      Contact( "CompALTA-MTA".FallaCompresor2 )
      wire#w4
      { S7_Templates := "SrcType := Int" } EQ_Contact(in1 := "DB-PrioridadesCmpAlta".Vcmp1, in2 := 2)
      wire#w5
      Contact( "DB-CompAltaDatos".Aut4 )
      Contact( "CompALTA-MTA".FallaCompresor4 )
      wire#w6
      { S7_Templates := "SrcType := Int" } EQ_Contact(in1 := "DB-PrioridadesCmpAlta".Vcmp4, in2 := 2)
   END_RUNG wire#w1
   RUNG wire#w4
      { S7_Templates := "SrcType := Int" } EQ_Contact(in1 := "DB-PrioridadesCmpAlta".Vcmp1, in2 := 1)
   END_RUNG wire#w5
   RUNG wire#w6
      { S7_Templates := "SrcType := Int" } EQ_Contact(in1 := "DB-PrioridadesCmpAlta".Vcmp4, in2 := 1)
   END_RUNG wire#w1
   RUNG wire#w5
      Contact( "DB-CompAltaDatos".Aut3 )
      Contact( "CompALTA-MTA".FallaCompresor3 )
      wire#w7
      { S7_Templates := "SrcType := Int" } EQ_Contact(in1 := "DB-PrioridadesCmpAlta".Vcmp3, in2 := 2)
   END_RUNG wire#w1
   RUNG wire#w7
      { S7_Templates := "SrcType := Int" } EQ_Contact(in1 := "DB-PrioridadesCmpAlta".Vcmp3, in2 := 1)
   END_RUNG wire#w1
   RUNG wire#w5
      Contact( "DB-CompAltaDatos".Aut2 )
      Contact( "CompALTA-MTA".FallaCompresor2 )
      wire#w8
      { S7_Templates := "SrcType := Int" } EQ_Contact(in1 := "DB-PrioridadesCmpAlta".Vcmp2, in2 := 2)
   END_RUNG wire#w1
   RUNG wire#w8
      { S7_Templates := "SrcType := Int" } EQ_Contact(in1 := "DB-PrioridadesCmpAlta".Vcmp2, in2 := 1)
   END_RUNG wire#w1
   RUNG wire#w3
      Contact( "DB-CompAltaDatos".Aut2 )
      Contact( "CompALTA-MTA".FallaCompresor2 )
      wire#w9
      { S7_Templates := "SrcType := Int" } EQ_Contact(in1 := "DB-PrioridadesCmpAlta".Vcmp2, in2 := 2)
      wire#w10
      Contact( "DB-CompAltaDatos".Aut4 )
      Contact( "CompALTA-MTA".FallaCompresor4 )
      wire#w11
      { S7_Templates := "SrcType := Int" } EQ_Contact(in1 := "DB-PrioridadesCmpAlta".Vcmp4, in2 := 2)
   END_RUNG wire#w1
   RUNG wire#w9
      { S7_Templates := "SrcType := Int" } EQ_Contact(in1 := "DB-PrioridadesCmpAlta".Vcmp2, in2 := 1)
   END_RUNG wire#w10
   RUNG wire#w11
      { S7_Templates := "SrcType := Int" } EQ_Contact(in1 := "DB-PrioridadesCmpAlta".Vcmp4, in2 := 1)
   END_RUNG wire#w1
   RUNG wire#w10
      Contact( "DB-CompAltaDatos".Aut3 )
      Contact( "CompALTA-MTA".FallaCompresor3 )
      wire#w12
      { S7_Templates := "SrcType := Int" } EQ_Contact(in1 := "DB-PrioridadesCmpAlta".Vcmp3, in2 := 2)
   END_RUNG wire#w1
   RUNG wire#w12
      { S7_Templates := "SrcType := Int" } EQ_Contact(in1 := "DB-PrioridadesCmpAlta".Vcmp3, in2 := 1)
   END_RUNG wire#w1
   RUNG wire#w3
      Contact( "DB-CompAltaDatos".Aut3 )
      Contact( "CompALTA-MTA".FallaCompresor3 )
      wire#w13
      { S7_Templates := "SrcType := Int" } EQ_Contact(in1 := "DB-PrioridadesCmpAlta".Vcmp3, in2 := 2)
      wire#w14
      Contact( "DB-CompAltaDatos".Aut4 )
      Contact( "CompALTA-MTA".FallaCompresor4 )
      wire#w15
      { S7_Templates := "SrcType := Int" } EQ_Contact(in1 := "DB-PrioridadesCmpAlta".Vcmp4, in2 := 2)
   END_RUNG wire#w1
   RUNG wire#w13
      { S7_Templates := "SrcType := Int" } EQ_Contact(in1 := "DB-PrioridadesCmpAlta".Vcmp3, in2 := 1)
   END_RUNG wire#w14
   RUNG wire#w15
      { S7_Templates := "SrcType := Int" } EQ_Contact(in1 := "DB-PrioridadesCmpAlta".Vcmp4, in2 := 1)
   END_RUNG wire#w1
   RUNG wire#powerrail
      { S7_Templates := "SrcType := Int" } EQ_Contact(in1 := "DB-PrioridadesCmpAlta".Vcmp5, in2 := 4)
      wire#w16
      Contact( "DB-CompAltaDatos".Aut1 )
      Contact( "CompALTA-MTA".FallaCompresor1 )
      wire#w17
      { S7_Templates := "SrcType := Int" } EQ_Contact(in1 := "DB-PrioridadesCmpAlta".Vcmp1, in2 := 3)
      wire#w18
      Contact( "DB-CompAltaDatos".Aut4 )
      Contact( "CompALTA-MTA".FallaCompresor4 )
      wire#w19
      { S7_Templates := "SrcType := Int" } EQ_Contact(in1 := "DB-PrioridadesCmpAlta".Vcmp4, in2 := 3)
      wire#w20
      Contact( "DB-CompAltaDatos".Aut2 )
      Contact( "CompALTA-MTA".FallaCompresor2 )
      wire#w21
      { S7_Templates := "SrcType := Int" } EQ_Contact(in1 := "DB-PrioridadesCmpAlta".Vcmp2, in2 := 3)
   END_RUNG wire#w1
   RUNG wire#w17
      { S7_Templates := "SrcType := Int" } EQ_Contact(in1 := "DB-PrioridadesCmpAlta".Vcmp1, in2 := 2)
   END_RUNG wire#w18
   RUNG wire#w17
      { S7_Templates := "SrcType := Int" } EQ_Contact(in1 := "DB-PrioridadesCmpAlta".Vcmp1, in2 := 1)
   END_RUNG wire#w18
   RUNG wire#w19
      { S7_Templates := "SrcType := Int" } EQ_Contact(in1 := "DB-PrioridadesCmpAlta".Vcmp4, in2 := 2)
   END_RUNG wire#w20
   RUNG wire#w19
      { S7_Templates := "SrcType := Int" } EQ_Contact(in1 := "DB-PrioridadesCmpAlta".Vcmp4, in2 := 1)
   END_RUNG wire#w20
   RUNG wire#w21
      { S7_Templates := "SrcType := Int" } EQ_Contact(in1 := "DB-PrioridadesCmpAlta".Vcmp2, in2 := 2)
   END_RUNG wire#w1
   RUNG wire#w21
      { S7_Templates := "SrcType := Int" } EQ_Contact(in1 := "DB-PrioridadesCmpAlta".Vcmp2, in2 := 1)
   END_RUNG wire#w1
   RUNG wire#w20
      Contact( "DB-CompAltaDatos".Aut4 )
      Contact( "CompALTA-MTA".FallaCompresor4 )
      wire#w22
      { S7_Templates := "SrcType := Int" } EQ_Contact(in1 := "DB-PrioridadesCmpAlta".Vcmp4, in2 := 3)
   END_RUNG wire#w1
   RUNG wire#w22
      { S7_Templates := "SrcType := Int" } EQ_Contact(in1 := "DB-PrioridadesCmpAlta".Vcmp4, in2 := 2)
   END_RUNG wire#w1
   RUNG wire#w22
      { S7_Templates := "SrcType := Int" } EQ_Contact(in1 := "DB-PrioridadesCmpAlta".Vcmp4, in2 := 1)
   END_RUNG wire#w1
   RUNG wire#w18
      Contact( "DB-CompAltaDatos".Aut3 )
      Contact( "CompALTA-MTA".FallaCompresor3 )
      wire#w23
      { S7_Templates := "SrcType := Int" } EQ_Contact(in1 := "DB-PrioridadesCmpAlta".Vcmp3, in2 := 3)
      wire#w24
      Contact( "DB-CompAltaDatos".Aut2 )
      Contact( "CompALTA-MTA".FallaCompresor2 )
      wire#w25
      { S7_Templates := "SrcType := Int" } EQ_Contact(in1 := "DB-PrioridadesCmpAlta".Vcmp2, in2 := 3)
   END_RUNG wire#w1
   RUNG wire#w23
      { S7_Templates := "SrcType := Int" } EQ_Contact(in1 := "DB-PrioridadesCmpAlta".Vcmp3, in2 := 2)
   END_RUNG wire#w24
   RUNG wire#w23
      { S7_Templates := "SrcType := Int" } EQ_Contact(in1 := "DB-PrioridadesCmpAlta".Vcmp3, in2 := 1)
   END_RUNG wire#w24
   RUNG wire#w25
      { S7_Templates := "SrcType := Int" } EQ_Contact(in1 := "DB-PrioridadesCmpAlta".Vcmp2, in2 := 2)
   END_RUNG wire#w1
   RUNG wire#w25
      { S7_Templates := "SrcType := Int" } EQ_Contact(in1 := "DB-PrioridadesCmpAlta".Vcmp2, in2 := 1)
   END_RUNG wire#w1
   RUNG wire#w16
      Contact( "DB-CompAltaDatos".Aut2 )
      Contact( "CompALTA-MTA".FallaCompresor2 )
      wire#w26
      { S7_Templates := "SrcType := Int" } EQ_Contact(in1 := "DB-PrioridadesCmpAlta".Vcmp2, in2 := 3)
      wire#w27
      Contact( "DB-CompAltaDatos".Aut4 )
      Contact( "CompALTA-MTA".FallaCompresor4 )
      wire#w28
      { S7_Templates := "SrcType := Int" } EQ_Contact(in1 := "DB-PrioridadesCmpAlta".Vcmp4, in2 := 3)
      wire#w29
      Contact( "DB-CompAltaDatos".Aut3 )
      Contact( "CompALTA-MTA".FallaCompresor3 )
      wire#w30
      { S7_Templates := "SrcType := Int" } EQ_Contact(in1 := "DB-PrioridadesCmpAlta".Vcmp3, in2 := 3)
   END_RUNG wire#w1
   RUNG wire#w26
      { S7_Templates := "SrcType := Int" } EQ_Contact(in1 := "DB-PrioridadesCmpAlta".Vcmp2, in2 := 2)
   END_RUNG wire#w27
   RUNG wire#w26
      { S7_Templates := "SrcType := Int" } EQ_Contact(in1 := "DB-PrioridadesCmpAlta".Vcmp2, in2 := 1)
   END_RUNG wire#w27
   RUNG wire#w28
      { S7_Templates := "SrcType := Int" } EQ_Contact(in1 := "DB-PrioridadesCmpAlta".Vcmp4, in2 := 2)
   END_RUNG wire#w29
   RUNG wire#w28
      { S7_Templates := "SrcType := Int" } EQ_Contact(in1 := "DB-PrioridadesCmpAlta".Vcmp4, in2 := 1)
   END_RUNG wire#w29
   RUNG wire#w30
      { S7_Templates := "SrcType := Int" } EQ_Contact(in1 := "DB-PrioridadesCmpAlta".Vcmp3, in2 := 2)
   END_RUNG wire#w1
   RUNG wire#w30
      { S7_Templates := "SrcType := Int" } EQ_Contact(in1 := "DB-PrioridadesCmpAlta".Vcmp3, in2 := 1)
   END_RUNG wire#w1
   RUNG wire#powerrail
      { S7_Templates := "SrcType := Int" } EQ_Contact(in1 := "DB-PrioridadesCmpAlta".Vcmp5, in2 := 5)
      Contact( "DB-CompAltaDatos".Aut1 )
      Contact( "CompALTA-MTA".FallaCompresor1 )
      Contact( "DB-CompAltaDatos".Aut2 )
      Contact( "CompALTA-MTA".FallaCompresor2 )
      Contact( "DB-CompAltaDatos".Aut3 )
      Contact( "CompALTA-MTA".FallaCompresor3 )
      Contact( "DB-CompAltaDatos".Aut4 )
      Contact( "CompALTA-MTA".FallaCompresor4 )
   END_RUNG wire#w1
   // the same network as SCL:
   IF (("DB-PrioridadesCmpAlta".Vcmp5 = 1) OR (("DB-PrioridadesCmpAlta".Vcmp5 = 2) AND (("DB-CompAltaDatos".Aut1 AND "CompALTA-MTA".FallaCompresor1 AND ("DB-PrioridadesCmpAlta".Vcmp1 = 1)) OR ("DB-CompAltaDatos".Aut2 AND "CompALTA-MTA".FallaCompresor2 AND ("DB-PrioridadesCmpAlta".Vcmp2 = 1)) OR ("DB-CompAltaDatos".Aut3 AND "CompALTA-MTA".FallaCompresor3 AND ("DB-PrioridadesCmpAlta".Vcmp3 = 1)) OR ("DB-CompAltaDatos".Aut4 AND "CompALTA-MTA".FallaCompresor4 AND ("DB-PrioridadesCmpAlta".Vcmp4 = 1)))) OR (("DB-PrioridadesCmpAlta".Vcmp5 = 3) AND (("DB-CompAltaDatos".Aut2 AND "CompALTA-MTA".FallaCompresor2 AND (("DB-PrioridadesCmpAlta".Vcmp1 = 2) OR ("DB-PrioridadesCmpAlta".Vcmp1 = 1)) AND (("DB-CompAltaDatos".Aut4 AND "CompALTA-MTA".FallaCompresor4 AND (("DB-PrioridadesCmpAlta".Vcmp4 = 2) OR ("DB-PrioridadesCmpAlta".Vcmp4 = 1))) OR ("DB-CompAltaDatos".Aut3 AND "CompALTA-MTA".FallaCompresor3 AND (("DB-PrioridadesCmpAlta".Vcmp3 = 2) OR ("DB-PrioridadesCmpAlta".Vcmp3 = 1))) OR ("DB-CompAltaDatos".Aut2 AND "CompALTA-MTA".FallaCompresor2 AND (("DB-PrioridadesCmpAlta".Vcmp2 = 2) OR ("DB-PrioridadesCmpAlta".Vcmp2 = 1))))) OR ("DB-CompAltaDatos".Aut2 AND "CompALTA-MTA".FallaCompresor2 AND (("DB-PrioridadesCmpAlta".Vcmp2 = 2) OR ("DB-PrioridadesCmpAlta".Vcmp2 = 1)) AND (("DB-CompAltaDatos".Aut4 AND "CompALTA-MTA".FallaCompresor4 AND (("DB-PrioridadesCmpAlta".Vcmp4 = 2) OR ("DB-PrioridadesCmpAlta".Vcmp4 = 1))) OR ("DB-CompAltaDatos".Aut3 AND "CompALTA-MTA".FallaCompresor3 AND (("DB-PrioridadesCmpAlta".Vcmp3 = 2) OR ("DB-PrioridadesCmpAlta".Vcmp3 = 1))))) OR ("DB-CompAltaDatos".Aut3 AND "CompALTA-MTA".FallaCompresor3 AND (("DB-PrioridadesCmpAlta".Vcmp3 = 2) OR ("DB-PrioridadesCmpAlta".Vcmp3 = 1)) AND "DB-CompAltaDatos".Aut4 AND "CompALTA-MTA".FallaCompresor4 AND (("DB-PrioridadesCmpAlta".Vcmp4 = 2) OR ("DB-PrioridadesCmpAlta".Vcmp4 = 1))))) OR (("DB-PrioridadesCmpAlta".Vcmp5 = 4) AND (("DB-CompAltaDatos".Aut1 AND "CompALTA-MTA".FallaCompresor1 AND (("DB-PrioridadesCmpAlta".Vcmp1 = 3) OR ("DB-PrioridadesCmpAlta".Vcmp1 = 2) OR ("DB-PrioridadesCmpAlta".Vcmp1 = 1)) AND (("DB-CompAltaDatos".Aut4 AND "CompALTA-MTA".FallaCompresor4 AND (("DB-PrioridadesCmpAlta".Vcmp4 = 3) OR ("DB-PrioridadesCmpAlta".Vcmp4 = 2) OR ("DB-PrioridadesCmpAlta".Vcmp4 = 1)) AND (("DB-CompAltaDatos".Aut2 AND "CompALTA-MTA".FallaCompresor2 AND (("DB-PrioridadesCmpAlta".Vcmp2 = 3) OR ("DB-PrioridadesCmpAlta".Vcmp2 = 2) OR ("DB-PrioridadesCmpAlta".Vcmp2 = 1))) OR ("DB-CompAltaDatos".Aut4 AND "CompALTA-MTA".FallaCompresor4 AND (("DB-PrioridadesCmpAlta".Vcmp4 = 3) OR ("DB-PrioridadesCmpAlta".Vcmp4 = 2) OR ("DB-PrioridadesCmpAlta".Vcmp4 = 1))))) OR ("DB-CompAltaDatos".Aut3 AND "CompALTA-MTA".FallaCompresor3 AND (("DB-PrioridadesCmpAlta".Vcmp3 = 3) OR ("DB-PrioridadesCmpAlta".Vcmp3 = 2) OR ("DB-PrioridadesCmpAlta".Vcmp3 = 1)) AND "DB-CompAltaDatos".Aut2 AND "CompALTA-MTA".FallaCompresor2 AND (("DB-PrioridadesCmpAlta".Vcmp2 = 3) OR ("DB-PrioridadesCmpAlta".Vcmp2 = 2) OR ("DB-PrioridadesCmpAlta".Vcmp2 = 1))))) OR ("DB-CompAltaDatos".Aut2 AND "CompALTA-MTA".FallaCompresor2 AND (("DB-PrioridadesCmpAlta".Vcmp2 = 3) OR ("DB-PrioridadesCmpAlta".Vcmp2 = 2) OR ("DB-PrioridadesCmpAlta".Vcmp2 = 1)) AND "DB-CompAltaDatos".Aut4 AND "CompALTA-MTA".FallaCompresor4 AND (("DB-PrioridadesCmpAlta".Vcmp4 = 3) OR ("DB-PrioridadesCmpAlta".Vcmp4 = 2) OR ("DB-PrioridadesCmpAlta".Vcmp4 = 1)) AND "DB-CompAltaDatos".Aut3 AND "CompALTA-MTA".FallaCompresor3 AND (("DB-PrioridadesCmpAlta".Vcmp3 = 3) OR ("DB-PrioridadesCmpAlta".Vcmp3 = 2) OR ("DB-PrioridadesCmpAlta".Vcmp3 = 1))))) OR (("DB-PrioridadesCmpAlta".Vcmp5 = 5) AND "DB-CompAltaDatos".Aut1 AND "CompALTA-MTA".FallaCompresor1 AND "DB-CompAltaDatos".Aut2 AND "CompALTA-MTA".FallaCompresor2 AND "DB-CompAltaDatos".Aut3 AND "CompALTA-MTA".FallaCompresor3 AND "DB-CompAltaDatos".Aut4 AND "CompALTA-MTA".FallaCompresor4)) AND "DB-CompAltaDatos".Aut5 AND NOT "CompALTA-MTA".FallaCompresor5 THEN
       "CompALTA-MTA".VRealCmp5 := 1;
   END_IF;
END_REGION
END_FUNCTION

FUNCTION "FlancosCmpAlta" : Void   // FC45, LAD
{ S7_Optimized_Access := 'FALSE' }
VERSION : 0.1
   VAR_TEMP   // added for the SCL form of the ladder/FBD networks
      _w1 : Bool;
      _w2 : Bool;
      _w3 : Bool;
      _w4 : Bool;
      _w5 : Bool;
      _w6 : Bool;
      _w7 : Bool;
      _s5time1 : S5Time;
   END_VAR
BEGIN

REGION Network 1
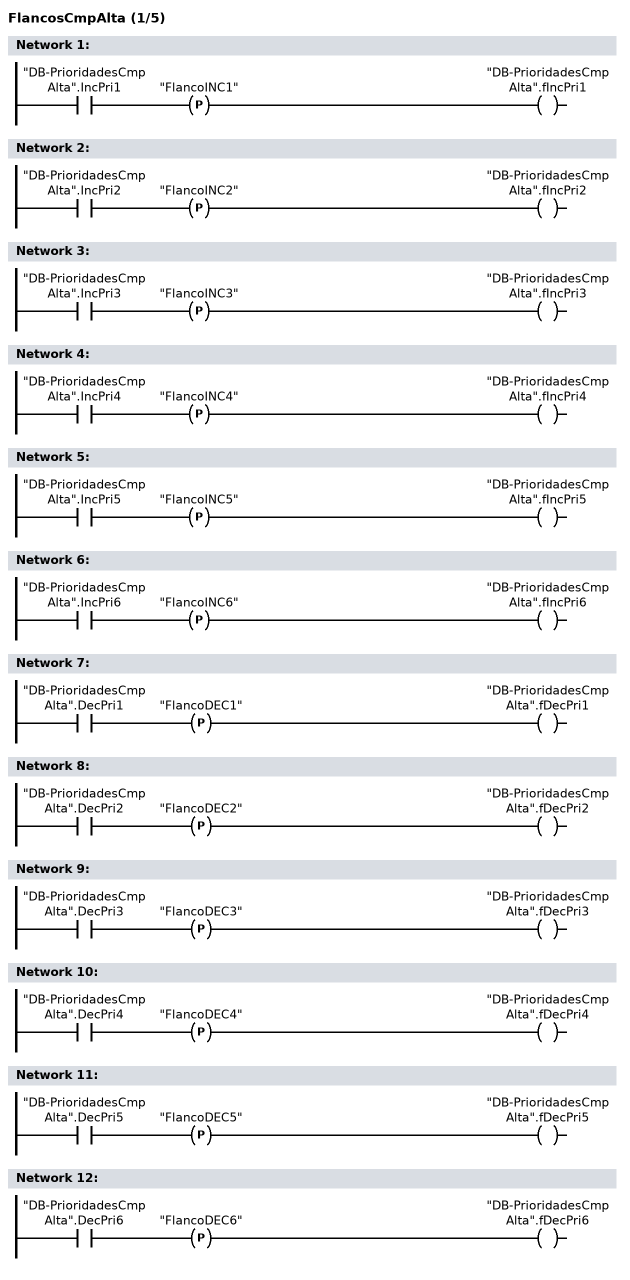
   RUNG wire#powerrail
      Contact( "DB-PrioridadesCmpAlta".IncPri1 )
      P_Trig( "FlancoINC1" )
      Coil( "DB-PrioridadesCmpAlta".fIncPri1 )
   END_RUNG
   // the same network as SCL:
   #_w1 := "DB-PrioridadesCmpAlta".IncPri1 AND NOT "FlancoINC1";   // rising edge
   "FlancoINC1" := "DB-PrioridadesCmpAlta".IncPri1;
   "DB-PrioridadesCmpAlta".fIncPri1 := #_w1;
END_REGION

REGION Network 2
   RUNG wire#powerrail
      Contact( "DB-PrioridadesCmpAlta".IncPri2 )
      P_Trig( "FlancoINC2" )
      Coil( "DB-PrioridadesCmpAlta".fIncPri2 )
   END_RUNG
   // the same network as SCL:
   #_w1 := "DB-PrioridadesCmpAlta".IncPri2 AND NOT "FlancoINC2";   // rising edge
   "FlancoINC2" := "DB-PrioridadesCmpAlta".IncPri2;
   "DB-PrioridadesCmpAlta".fIncPri2 := #_w1;
END_REGION

REGION Network 3
   RUNG wire#powerrail
      Contact( "DB-PrioridadesCmpAlta".IncPri3 )
      P_Trig( "FlancoINC3" )
      Coil( "DB-PrioridadesCmpAlta".fIncPri3 )
   END_RUNG
   // the same network as SCL:
   #_w1 := "DB-PrioridadesCmpAlta".IncPri3 AND NOT "FlancoINC3";   // rising edge
   "FlancoINC3" := "DB-PrioridadesCmpAlta".IncPri3;
   "DB-PrioridadesCmpAlta".fIncPri3 := #_w1;
END_REGION

REGION Network 4
   RUNG wire#powerrail
      Contact( "DB-PrioridadesCmpAlta".IncPri4 )
      P_Trig( "FlancoINC4" )
      Coil( "DB-PrioridadesCmpAlta".fIncPri4 )
   END_RUNG
   // the same network as SCL:
   #_w1 := "DB-PrioridadesCmpAlta".IncPri4 AND NOT "FlancoINC4";   // rising edge
   "FlancoINC4" := "DB-PrioridadesCmpAlta".IncPri4;
   "DB-PrioridadesCmpAlta".fIncPri4 := #_w1;
END_REGION

REGION Network 5
   RUNG wire#powerrail
      Contact( "DB-PrioridadesCmpAlta".IncPri5 )
      P_Trig( "FlancoINC5" )
      Coil( "DB-PrioridadesCmpAlta".fIncPri5 )
   END_RUNG
   // the same network as SCL:
   #_w1 := "DB-PrioridadesCmpAlta".IncPri5 AND NOT "FlancoINC5";   // rising edge
   "FlancoINC5" := "DB-PrioridadesCmpAlta".IncPri5;
   "DB-PrioridadesCmpAlta".fIncPri5 := #_w1;
END_REGION

REGION Network 6
   RUNG wire#powerrail
      Contact( "DB-PrioridadesCmpAlta".IncPri6 )
      P_Trig( "FlancoINC6" )
      Coil( "DB-PrioridadesCmpAlta".fIncPri6 )
   END_RUNG
   // the same network as SCL:
   #_w1 := "DB-PrioridadesCmpAlta".IncPri6 AND NOT "FlancoINC6";   // rising edge
   "FlancoINC6" := "DB-PrioridadesCmpAlta".IncPri6;
   "DB-PrioridadesCmpAlta".fIncPri6 := #_w1;
END_REGION

REGION Network 7
   RUNG wire#powerrail
      Contact( "DB-PrioridadesCmpAlta".DecPri1 )
      P_Trig( "FlancoDEC1" )
      Coil( "DB-PrioridadesCmpAlta".fDecPri1 )
   END_RUNG
   // the same network as SCL:
   #_w1 := "DB-PrioridadesCmpAlta".DecPri1 AND NOT "FlancoDEC1";   // rising edge
   "FlancoDEC1" := "DB-PrioridadesCmpAlta".DecPri1;
   "DB-PrioridadesCmpAlta".fDecPri1 := #_w1;
END_REGION

REGION Network 8
   RUNG wire#powerrail
      Contact( "DB-PrioridadesCmpAlta".DecPri2 )
      P_Trig( "FlancoDEC2" )
      Coil( "DB-PrioridadesCmpAlta".fDecPri2 )
   END_RUNG
   // the same network as SCL:
   #_w1 := "DB-PrioridadesCmpAlta".DecPri2 AND NOT "FlancoDEC2";   // rising edge
   "FlancoDEC2" := "DB-PrioridadesCmpAlta".DecPri2;
   "DB-PrioridadesCmpAlta".fDecPri2 := #_w1;
END_REGION

REGION Network 9
   RUNG wire#powerrail
      Contact( "DB-PrioridadesCmpAlta".DecPri3 )
      P_Trig( "FlancoDEC3" )
      Coil( "DB-PrioridadesCmpAlta".fDecPri3 )
   END_RUNG
   // the same network as SCL:
   #_w1 := "DB-PrioridadesCmpAlta".DecPri3 AND NOT "FlancoDEC3";   // rising edge
   "FlancoDEC3" := "DB-PrioridadesCmpAlta".DecPri3;
   "DB-PrioridadesCmpAlta".fDecPri3 := #_w1;
END_REGION

REGION Network 10
   RUNG wire#powerrail
      Contact( "DB-PrioridadesCmpAlta".DecPri4 )
      P_Trig( "FlancoDEC4" )
      Coil( "DB-PrioridadesCmpAlta".fDecPri4 )
   END_RUNG
   // the same network as SCL:
   #_w1 := "DB-PrioridadesCmpAlta".DecPri4 AND NOT "FlancoDEC4";   // rising edge
   "FlancoDEC4" := "DB-PrioridadesCmpAlta".DecPri4;
   "DB-PrioridadesCmpAlta".fDecPri4 := #_w1;
END_REGION

REGION Network 11
   RUNG wire#powerrail
      Contact( "DB-PrioridadesCmpAlta".DecPri5 )
      P_Trig( "FlancoDEC5" )
      Coil( "DB-PrioridadesCmpAlta".fDecPri5 )
   END_RUNG
   // the same network as SCL:
   #_w1 := "DB-PrioridadesCmpAlta".DecPri5 AND NOT "FlancoDEC5";   // rising edge
   "FlancoDEC5" := "DB-PrioridadesCmpAlta".DecPri5;
   "DB-PrioridadesCmpAlta".fDecPri5 := #_w1;
END_REGION

REGION Network 12
   RUNG wire#powerrail
      Contact( "DB-PrioridadesCmpAlta".DecPri6 )
      P_Trig( "FlancoDEC6" )
      Coil( "DB-PrioridadesCmpAlta".fDecPri6 )
   END_RUNG
   // the same network as SCL:
   #_w1 := "DB-PrioridadesCmpAlta".DecPri6 AND NOT "FlancoDEC6";   // rising edge
   "FlancoDEC6" := "DB-PrioridadesCmpAlta".DecPri6;
   "DB-PrioridadesCmpAlta".fDecPri6 := #_w1;
END_REGION

REGION Network 13
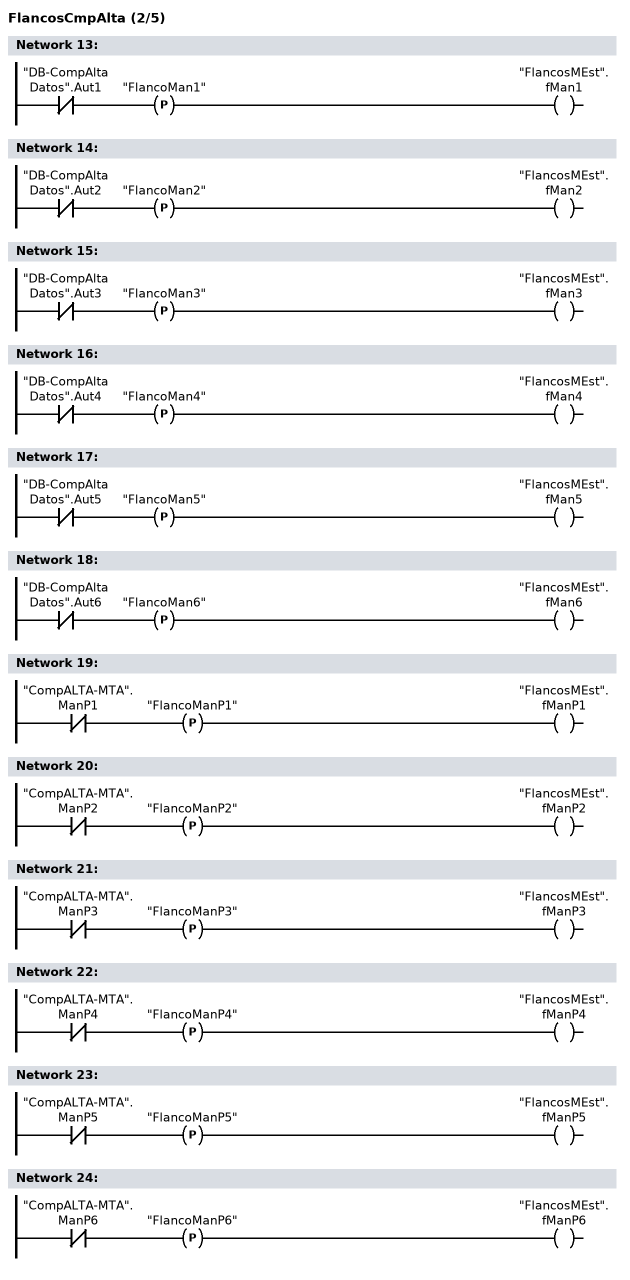
   RUNG wire#powerrail
      I_Contact( "DB-CompAltaDatos".Aut1 )
      P_Trig( "FlancoMan1" )
      Coil( "FlancosMEst".fMan1 )
   END_RUNG
   // the same network as SCL:
   #_w1 := NOT "DB-CompAltaDatos".Aut1 AND NOT "FlancoMan1";   // rising edge
   "FlancoMan1" := NOT "DB-CompAltaDatos".Aut1;
   "FlancosMEst".fMan1 := #_w1;
END_REGION

REGION Network 14
   RUNG wire#powerrail
      I_Contact( "DB-CompAltaDatos".Aut2 )
      P_Trig( "FlancoMan2" )
      Coil( "FlancosMEst".fMan2 )
   END_RUNG
   // the same network as SCL:
   #_w1 := NOT "DB-CompAltaDatos".Aut2 AND NOT "FlancoMan2";   // rising edge
   "FlancoMan2" := NOT "DB-CompAltaDatos".Aut2;
   "FlancosMEst".fMan2 := #_w1;
END_REGION

REGION Network 15
   RUNG wire#powerrail
      I_Contact( "DB-CompAltaDatos".Aut3 )
      P_Trig( "FlancoMan3" )
      Coil( "FlancosMEst".fMan3 )
   END_RUNG
   // the same network as SCL:
   #_w1 := NOT "DB-CompAltaDatos".Aut3 AND NOT "FlancoMan3";   // rising edge
   "FlancoMan3" := NOT "DB-CompAltaDatos".Aut3;
   "FlancosMEst".fMan3 := #_w1;
END_REGION

REGION Network 16
   RUNG wire#powerrail
      I_Contact( "DB-CompAltaDatos".Aut4 )
      P_Trig( "FlancoMan4" )
      Coil( "FlancosMEst".fMan4 )
   END_RUNG
   // the same network as SCL:
   #_w1 := NOT "DB-CompAltaDatos".Aut4 AND NOT "FlancoMan4";   // rising edge
   "FlancoMan4" := NOT "DB-CompAltaDatos".Aut4;
   "FlancosMEst".fMan4 := #_w1;
END_REGION

REGION Network 17
   RUNG wire#powerrail
      I_Contact( "DB-CompAltaDatos".Aut5 )
      P_Trig( "FlancoMan5" )
      Coil( "FlancosMEst".fMan5 )
   END_RUNG
   // the same network as SCL:
   #_w1 := NOT "DB-CompAltaDatos".Aut5 AND NOT "FlancoMan5";   // rising edge
   "FlancoMan5" := NOT "DB-CompAltaDatos".Aut5;
   "FlancosMEst".fMan5 := #_w1;
END_REGION

REGION Network 18
   RUNG wire#powerrail
      I_Contact( "DB-CompAltaDatos".Aut6 )
      P_Trig( "FlancoMan6" )
      Coil( "FlancosMEst".fMan6 )
   END_RUNG
   // the same network as SCL:
   #_w1 := NOT "DB-CompAltaDatos".Aut6 AND NOT "FlancoMan6";   // rising edge
   "FlancoMan6" := NOT "DB-CompAltaDatos".Aut6;
   "FlancosMEst".fMan6 := #_w1;
END_REGION

REGION Network 19
   RUNG wire#powerrail
      I_Contact( "CompALTA-MTA".ManP1 )
      P_Trig( "FlancoManP1" )
      Coil( "FlancosMEst".fManP1 )
   END_RUNG
   // the same network as SCL:
   #_w1 := NOT "CompALTA-MTA".ManP1 AND NOT "FlancoManP1";   // rising edge
   "FlancoManP1" := NOT "CompALTA-MTA".ManP1;
   "FlancosMEst".fManP1 := #_w1;
END_REGION

REGION Network 20
   RUNG wire#powerrail
      I_Contact( "CompALTA-MTA".ManP2 )
      P_Trig( "FlancoManP2" )
      Coil( "FlancosMEst".fManP2 )
   END_RUNG
   // the same network as SCL:
   #_w1 := NOT "CompALTA-MTA".ManP2 AND NOT "FlancoManP2";   // rising edge
   "FlancoManP2" := NOT "CompALTA-MTA".ManP2;
   "FlancosMEst".fManP2 := #_w1;
END_REGION

REGION Network 21
   RUNG wire#powerrail
      I_Contact( "CompALTA-MTA".ManP3 )
      P_Trig( "FlancoManP3" )
      Coil( "FlancosMEst".fManP3 )
   END_RUNG
   // the same network as SCL:
   #_w1 := NOT "CompALTA-MTA".ManP3 AND NOT "FlancoManP3";   // rising edge
   "FlancoManP3" := NOT "CompALTA-MTA".ManP3;
   "FlancosMEst".fManP3 := #_w1;
END_REGION

REGION Network 22
   RUNG wire#powerrail
      I_Contact( "CompALTA-MTA".ManP4 )
      P_Trig( "FlancoManP4" )
      Coil( "FlancosMEst".fManP4 )
   END_RUNG
   // the same network as SCL:
   #_w1 := NOT "CompALTA-MTA".ManP4 AND NOT "FlancoManP4";   // rising edge
   "FlancoManP4" := NOT "CompALTA-MTA".ManP4;
   "FlancosMEst".fManP4 := #_w1;
END_REGION

REGION Network 23
   RUNG wire#powerrail
      I_Contact( "CompALTA-MTA".ManP5 )
      P_Trig( "FlancoManP5" )
      Coil( "FlancosMEst".fManP5 )
   END_RUNG
   // the same network as SCL:
   #_w1 := NOT "CompALTA-MTA".ManP5 AND NOT "FlancoManP5";   // rising edge
   "FlancoManP5" := NOT "CompALTA-MTA".ManP5;
   "FlancosMEst".fManP5 := #_w1;
END_REGION

REGION Network 24
   RUNG wire#powerrail
      I_Contact( "CompALTA-MTA".ManP6 )
      P_Trig( "FlancoManP6" )
      Coil( "FlancosMEst".fManP6 )
   END_RUNG
   // the same network as SCL:
   #_w1 := NOT "CompALTA-MTA".ManP6 AND NOT "FlancoManP6";   // rising edge
   "FlancoManP6" := NOT "CompALTA-MTA".ManP6;
   "FlancosMEst".fManP6 := #_w1;
END_REGION

REGION Network 25
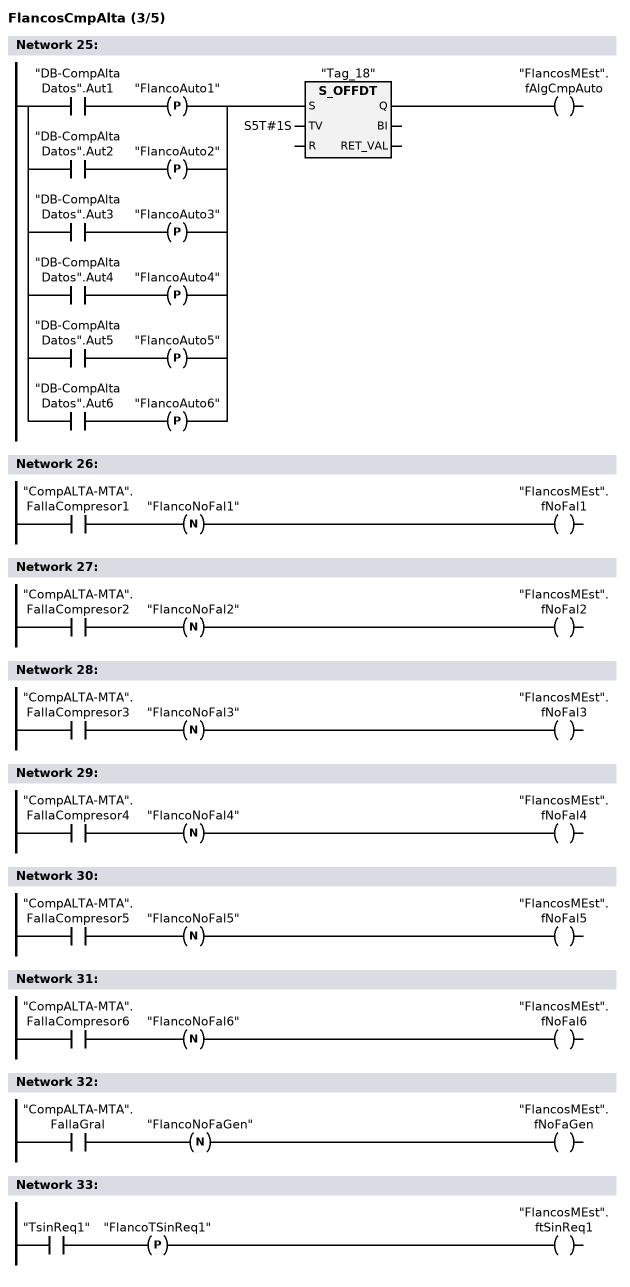
   RUNG wire#powerrail
      Contact( "DB-CompAltaDatos".Aut1 )
      P_Trig( "FlancoAuto1" )
      wire#w1
      S_OFFDT(T_NO := "Tag_18", TV := S5T#1S, R :=, BI =>, RET_VAL =>)
      Coil( "FlancosMEst".fAlgCmpAuto )
   END_RUNG
   RUNG wire#powerrail
      Contact( "DB-CompAltaDatos".Aut2 )
      P_Trig( "FlancoAuto2" )
   END_RUNG wire#w1
   RUNG wire#powerrail
      Contact( "DB-CompAltaDatos".Aut3 )
      P_Trig( "FlancoAuto3" )
   END_RUNG wire#w1
   RUNG wire#powerrail
      Contact( "DB-CompAltaDatos".Aut4 )
      P_Trig( "FlancoAuto4" )
   END_RUNG wire#w1
   RUNG wire#powerrail
      Contact( "DB-CompAltaDatos".Aut5 )
      P_Trig( "FlancoAuto5" )
   END_RUNG wire#w1
   RUNG wire#powerrail
      Contact( "DB-CompAltaDatos".Aut6 )
      P_Trig( "FlancoAuto6" )
   END_RUNG wire#w1
   // the same network as SCL:
   #_w1 := "DB-CompAltaDatos".Aut1 AND NOT "FlancoAuto1";   // rising edge
   "FlancoAuto1" := "DB-CompAltaDatos".Aut1;
   #_w2 := "DB-CompAltaDatos".Aut2 AND NOT "FlancoAuto2";   // rising edge
   "FlancoAuto2" := "DB-CompAltaDatos".Aut2;
   #_w3 := "DB-CompAltaDatos".Aut3 AND NOT "FlancoAuto3";   // rising edge
   "FlancoAuto3" := "DB-CompAltaDatos".Aut3;
   #_w4 := "DB-CompAltaDatos".Aut4 AND NOT "FlancoAuto4";   // rising edge
   "FlancoAuto4" := "DB-CompAltaDatos".Aut4;
   #_w5 := "DB-CompAltaDatos".Aut5 AND NOT "FlancoAuto5";   // rising edge
   "FlancoAuto5" := "DB-CompAltaDatos".Aut5;
   #_w6 := "DB-CompAltaDatos".Aut6 AND NOT "FlancoAuto6";   // rising edge
   "FlancoAuto6" := "DB-CompAltaDatos".Aut6;
   #_s5time1 := S_OFFDT(T_NO := "Tag_18",
                        S := #_w1 OR #_w2 OR #_w3 OR #_w4 OR #_w5 OR #_w6,
                        TV := S5T#1S,
                        Q => #_w7);
   "FlancosMEst".fAlgCmpAuto := #_w7;
END_REGION

REGION Network 26
   RUNG wire#powerrail
      Contact( "CompALTA-MTA".FallaCompresor1 )
      N_Trig( "FlancoNoFal1" )
      Coil( "FlancosMEst".fNoFal1 )
   END_RUNG
   // the same network as SCL:
   #_w1 := NOT "CompALTA-MTA".FallaCompresor1 AND "FlancoNoFal1";   // falling edge
   "FlancoNoFal1" := "CompALTA-MTA".FallaCompresor1;
   "FlancosMEst".fNoFal1 := #_w1;
END_REGION

REGION Network 27
   RUNG wire#powerrail
      Contact( "CompALTA-MTA".FallaCompresor2 )
      N_Trig( "FlancoNoFal2" )
      Coil( "FlancosMEst".fNoFal2 )
   END_RUNG
   // the same network as SCL:
   #_w1 := NOT "CompALTA-MTA".FallaCompresor2 AND "FlancoNoFal2";   // falling edge
   "FlancoNoFal2" := "CompALTA-MTA".FallaCompresor2;
   "FlancosMEst".fNoFal2 := #_w1;
END_REGION

REGION Network 28
   RUNG wire#powerrail
      Contact( "CompALTA-MTA".FallaCompresor3 )
      N_Trig( "FlancoNoFal3" )
      Coil( "FlancosMEst".fNoFal3 )
   END_RUNG
   // the same network as SCL:
   #_w1 := NOT "CompALTA-MTA".FallaCompresor3 AND "FlancoNoFal3";   // falling edge
   "FlancoNoFal3" := "CompALTA-MTA".FallaCompresor3;
   "FlancosMEst".fNoFal3 := #_w1;
END_REGION

REGION Network 29
   RUNG wire#powerrail
      Contact( "CompALTA-MTA".FallaCompresor4 )
      N_Trig( "FlancoNoFal4" )
      Coil( "FlancosMEst".fNoFal4 )
   END_RUNG
   // the same network as SCL:
   #_w1 := NOT "CompALTA-MTA".FallaCompresor4 AND "FlancoNoFal4";   // falling edge
   "FlancoNoFal4" := "CompALTA-MTA".FallaCompresor4;
   "FlancosMEst".fNoFal4 := #_w1;
END_REGION

REGION Network 30
   RUNG wire#powerrail
      Contact( "CompALTA-MTA".FallaCompresor5 )
      N_Trig( "FlancoNoFal5" )
      Coil( "FlancosMEst".fNoFal5 )
   END_RUNG
   // the same network as SCL:
   #_w1 := NOT "CompALTA-MTA".FallaCompresor5 AND "FlancoNoFal5";   // falling edge
   "FlancoNoFal5" := "CompALTA-MTA".FallaCompresor5;
   "FlancosMEst".fNoFal5 := #_w1;
END_REGION

REGION Network 31
   RUNG wire#powerrail
      Contact( "CompALTA-MTA".FallaCompresor6 )
      N_Trig( "FlancoNoFal6" )
      Coil( "FlancosMEst".fNoFal6 )
   END_RUNG
   // the same network as SCL:
   #_w1 := NOT "CompALTA-MTA".FallaCompresor6 AND "FlancoNoFal6";   // falling edge
   "FlancoNoFal6" := "CompALTA-MTA".FallaCompresor6;
   "FlancosMEst".fNoFal6 := #_w1;
END_REGION

REGION Network 32
   RUNG wire#powerrail
      Contact( "CompALTA-MTA".FallaGral )
      N_Trig( "FlancoNoFaGen" )
      Coil( "FlancosMEst".fNoFaGen )
   END_RUNG
   // the same network as SCL:
   #_w1 := NOT "CompALTA-MTA".FallaGral AND "FlancoNoFaGen";   // falling edge
   "FlancoNoFaGen" := "CompALTA-MTA".FallaGral;
   "FlancosMEst".fNoFaGen := #_w1;
END_REGION

REGION Network 33
   RUNG wire#powerrail
      Contact( "TsinReq1" )
      P_Trig( "FlancoTSinReq1" )
      Coil( "FlancosMEst".ftSinReq1 )
   END_RUNG
   // the same network as SCL:
   #_w1 := "TsinReq1" AND NOT "FlancoTSinReq1";   // rising edge
   "FlancoTSinReq1" := "TsinReq1";
   "FlancosMEst".ftSinReq1 := #_w1;
END_REGION

REGION Network 34
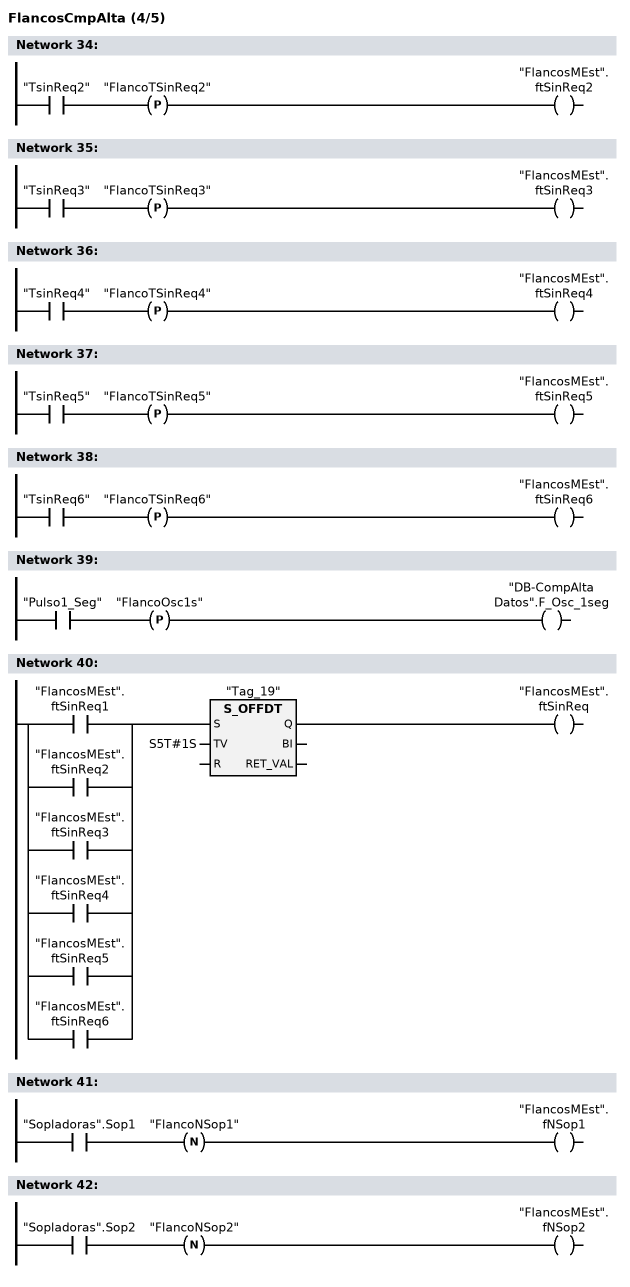
   RUNG wire#powerrail
      Contact( "TsinReq2" )
      P_Trig( "FlancoTSinReq2" )
      Coil( "FlancosMEst".ftSinReq2 )
   END_RUNG
   // the same network as SCL:
   #_w1 := "TsinReq2" AND NOT "FlancoTSinReq2";   // rising edge
   "FlancoTSinReq2" := "TsinReq2";
   "FlancosMEst".ftSinReq2 := #_w1;
END_REGION

REGION Network 35
   RUNG wire#powerrail
      Contact( "TsinReq3" )
      P_Trig( "FlancoTSinReq3" )
      Coil( "FlancosMEst".ftSinReq3 )
   END_RUNG
   // the same network as SCL:
   #_w1 := "TsinReq3" AND NOT "FlancoTSinReq3";   // rising edge
   "FlancoTSinReq3" := "TsinReq3";
   "FlancosMEst".ftSinReq3 := #_w1;
END_REGION

REGION Network 36
   RUNG wire#powerrail
      Contact( "TsinReq4" )
      P_Trig( "FlancoTSinReq4" )
      Coil( "FlancosMEst".ftSinReq4 )
   END_RUNG
   // the same network as SCL:
   #_w1 := "TsinReq4" AND NOT "FlancoTSinReq4";   // rising edge
   "FlancoTSinReq4" := "TsinReq4";
   "FlancosMEst".ftSinReq4 := #_w1;
END_REGION

REGION Network 37
   RUNG wire#powerrail
      Contact( "TsinReq5" )
      P_Trig( "FlancoTSinReq5" )
      Coil( "FlancosMEst".ftSinReq5 )
   END_RUNG
   // the same network as SCL:
   #_w1 := "TsinReq5" AND NOT "FlancoTSinReq5";   // rising edge
   "FlancoTSinReq5" := "TsinReq5";
   "FlancosMEst".ftSinReq5 := #_w1;
END_REGION

REGION Network 38
   RUNG wire#powerrail
      Contact( "TsinReq6" )
      P_Trig( "FlancoTSinReq6" )
      Coil( "FlancosMEst".ftSinReq6 )
   END_RUNG
   // the same network as SCL:
   #_w1 := "TsinReq6" AND NOT "FlancoTSinReq6";   // rising edge
   "FlancoTSinReq6" := "TsinReq6";
   "FlancosMEst".ftSinReq6 := #_w1;
END_REGION

REGION Network 39
   RUNG wire#powerrail
      Contact( "Pulso1_Seg" )
      P_Trig( "FlancoOsc1s" )
      Coil( "DB-CompAltaDatos".F_Osc_1seg )
   END_RUNG
   // the same network as SCL:
   #_w1 := "Pulso1_Seg" AND NOT "FlancoOsc1s";   // rising edge
   "FlancoOsc1s" := "Pulso1_Seg";
   "DB-CompAltaDatos".F_Osc_1seg := #_w1;
END_REGION

REGION Network 40
   RUNG wire#powerrail
      Contact( "FlancosMEst".ftSinReq1 )
      wire#w1
      S_OFFDT(T_NO := "Tag_19", TV := S5T#1S, R :=, BI =>, RET_VAL =>)
      Coil( "FlancosMEst".ftSinReq )
   END_RUNG
   RUNG wire#powerrail
      Contact( "FlancosMEst".ftSinReq2 )
   END_RUNG wire#w1
   RUNG wire#powerrail
      Contact( "FlancosMEst".ftSinReq3 )
   END_RUNG wire#w1
   RUNG wire#powerrail
      Contact( "FlancosMEst".ftSinReq4 )
   END_RUNG wire#w1
   RUNG wire#powerrail
      Contact( "FlancosMEst".ftSinReq5 )
   END_RUNG wire#w1
   RUNG wire#powerrail
      Contact( "FlancosMEst".ftSinReq6 )
   END_RUNG wire#w1
   // the same network as SCL:
   #_s5time1 := S_OFFDT(T_NO := "Tag_19",
                        S := "FlancosMEst".ftSinReq1 OR "FlancosMEst".ftSinReq2 OR "FlancosMEst".ftSinReq3 OR "FlancosMEst".ftSinReq4 OR "FlancosMEst".ftSinReq5 OR "FlancosMEst".ftSinReq6,
                        TV := S5T#1S,
                        Q => #_w1);
   "FlancosMEst".ftSinReq := #_w1;
END_REGION

REGION Network 41
   RUNG wire#powerrail
      Contact( "Sopladoras".Sop1 )
      N_Trig( "FlancoNSop1" )
      Coil( "FlancosMEst".fNSop1 )
   END_RUNG
   // the same network as SCL:
   #_w1 := NOT "Sopladoras".Sop1 AND "FlancoNSop1";   // falling edge
   "FlancoNSop1" := "Sopladoras".Sop1;
   "FlancosMEst".fNSop1 := #_w1;
END_REGION

REGION Network 42
   RUNG wire#powerrail
      Contact( "Sopladoras".Sop2 )
      N_Trig( "FlancoNSop2" )
      Coil( "FlancosMEst".fNSop2 )
   END_RUNG
   // the same network as SCL:
   #_w1 := NOT "Sopladoras".Sop2 AND "FlancoNSop2";   // falling edge
   "FlancoNSop2" := "Sopladoras".Sop2;
   "FlancosMEst".fNSop2 := #_w1;
END_REGION

REGION Network 43
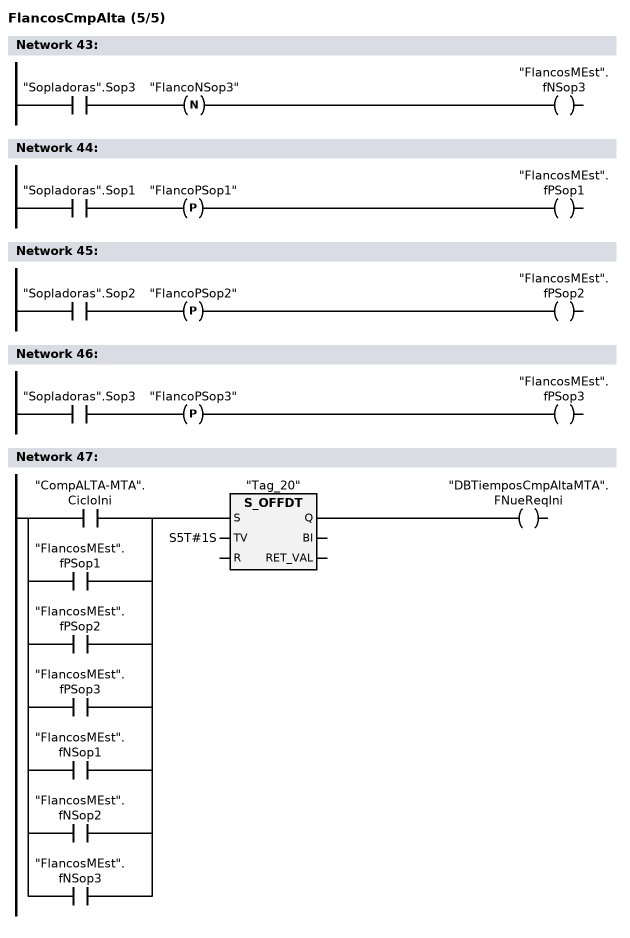
   RUNG wire#powerrail
      Contact( "Sopladoras".Sop3 )
      N_Trig( "FlancoNSop3" )
      Coil( "FlancosMEst".fNSop3 )
   END_RUNG
   // the same network as SCL:
   #_w1 := NOT "Sopladoras".Sop3 AND "FlancoNSop3";   // falling edge
   "FlancoNSop3" := "Sopladoras".Sop3;
   "FlancosMEst".fNSop3 := #_w1;
END_REGION

REGION Network 44
   RUNG wire#powerrail
      Contact( "Sopladoras".Sop1 )
      P_Trig( "FlancoPSop1" )
      Coil( "FlancosMEst".fPSop1 )
   END_RUNG
   // the same network as SCL:
   #_w1 := "Sopladoras".Sop1 AND NOT "FlancoPSop1";   // rising edge
   "FlancoPSop1" := "Sopladoras".Sop1;
   "FlancosMEst".fPSop1 := #_w1;
END_REGION

REGION Network 45
   RUNG wire#powerrail
      Contact( "Sopladoras".Sop2 )
      P_Trig( "FlancoPSop2" )
      Coil( "FlancosMEst".fPSop2 )
   END_RUNG
   // the same network as SCL:
   #_w1 := "Sopladoras".Sop2 AND NOT "FlancoPSop2";   // rising edge
   "FlancoPSop2" := "Sopladoras".Sop2;
   "FlancosMEst".fPSop2 := #_w1;
END_REGION

REGION Network 46
   RUNG wire#powerrail
      Contact( "Sopladoras".Sop3 )
      P_Trig( "FlancoPSop3" )
      Coil( "FlancosMEst".fPSop3 )
   END_RUNG
   // the same network as SCL:
   #_w1 := "Sopladoras".Sop3 AND NOT "FlancoPSop3";   // rising edge
   "FlancoPSop3" := "Sopladoras".Sop3;
   "FlancosMEst".fPSop3 := #_w1;
END_REGION

